        rgtPlate[1].tData.rgtCap[0].tFlag.tSelvedgeMachine.dDoneTrim1OpSide := 3, rgtPlate[1].tData.rgtCap[0].tFlag.tSelvedgeMachine.dDoneTrim2OppOpSide := 1, rgtPlate[1].tData.rgtCap[0].tFlag.tSelvedgeMachine.dDoneTrim3OppOpSide := 3, rgtPlate[2].tTracking.dPosition_cmm := 2104636, rgtPlate[2].tTracking.dPositionHead_cmm := 2234636, rgtPlate[2].tTracking.dPositionTail_cmm := 1974636, rgtPlate[2].tTracking.dLength_cmm := 260000, rgtPlate[2].tTracking.dIndexConvHead := 7, rgtPlate[2].tTracking.dIndexCapInConvHead := 2, rgtPlate[2].tTracking.dIndexConvTail := 6, rgtPlate[2].tTracking.dIndexCapInConvTail := 2, rgtPlate[2].tTracking.dLastConv := 6, rgtPlate[2].tTracking.dLastConvTail := 6, rgtPlate[2].tData.dLength_cmm := 260000, rgtPlate[2].tData.dTotalCaps := 1, rgtPlate[2].tData.rgtCap[0].dID := 4255236, rgtPlate[2].tData.rgtCap[0].dLength_cmm := 260000, rgtPlate[2].tData.rgtCap[0].dWidth_cmm := 360000, rgtPlate[2].tData.rgtCap[0].dThickness_cmm := 600, rgtPlate[2].tData.rgtCap[0].dFormat := 3, rgtPlate[2].tData.rgtCap[0].dNumLites := 2, rgtPlate[2].tData.rgtCap[0].dConvTotLength_cmm := 260000, rgtPlate[2].tData.rgtCap[0].dMinWidth_cmm := 360000, rgtPlate[2].tData.rgtCap[0].dMaxWidth_cmm := 360000, rgtPlate[2].tData.rgtCap[0].dGrossWidth_cmm := 377300, rgtPlate[2].tData.rgtCap[0].dDEdgeOpSide_cmm := 5000, rgtPlate[2].tData.rgtCap[0].dDEdgeOppOpSide_cmm := 5000, rgtPlate[2].tData.rgtCap[0].dCutWander_cmm := -3930, rgtPlate[2].tData.rgtCap[0].dNetWander_cmm := -6230, rgtPlate[2].tData.rgtCap[0].rgtLite[0].dID := 4255237, rgtPlate[2].tData.rgtCap[0].rgtLite[0].dProductionID := 1029, rgtPlate[2].tData.rgtCap[0].rgtLite[0].dQualityID := 10, rgtPlate[2].tData.rgtCap[0].rgtLite[0].dWidth_cmm := 180000, rgtPlate[2].tData.rgtCap[0].rgtLite[0].dBarycenter_cmm := -93930, rgtPlate[2].tData.rgtCap[0].rgtLite[1].dID := 4255238, rgtPlate[2].tData.rgtCap[0].rgtLite[1].dProductionID := 1029, rgtPlate[2].tData.rgtCap[0].rgtLite[1].dQualityID := 10, rgtPlate[2].tData.rgtCap[0].rgtLite[1].dWidth_cmm := 180000, rgtPlate[2].tData.rgtCap[0].rgtLite[1].dBarycenter_cmm := 86070, rgtPlate[2].tData.rgtCap[0].tFlag.xByYCut2 := 1, rgtPlate[2].tData.rgtCap[0].tFlag.xTrim2OpSide := 1, rgtPlate[2].tData.rgtCap[0].tFlag.xTrim1OpSide := 1, rgtPlate[2].tData.rgtCap[0].tFlag.xTrim1OppOpSide := 1, rgtPlate[2].tData.rgtCap[0].tFlag.xTrim2OppOpSide := 1, rgtPlate[2].tData.rgtCap[0].tFlag.rgxIntCut := 1, rgtPlate[2].tData.rgtCap[0].tFlag.xOptSelvedgeSel := 1, rgtPlate[2].tData.rgtCap[0].tFlag.xOptSplitBarSel := 1, rgtPlate[2].tData.rgtCap[0].tFlag.xOptSepRollSel := 1, rgtPlate[2].tData.rgtCap[0].tFlag.rgxXCutDoneHead := 2, rgtPlate[2].tData.rgtCap[0].tFlag.rgxXCutDoneTail := 2, rgtPlate[2].tData.rgtCap[0].tFlag.rgxYCutHeadDone := 835, rgtPlate[2].tData.rgtCap[0].tFlag.tSelvedgeMachine.dReqTrim2OpSide := 1, rgtPlate[2].tData.rgtCap[0].tFlag.tSelvedgeMachine.dReqTrim1OpSide := 3, rgtPlate[2].tData.rgtCap[0].tFlag.tSelvedgeMachine.dReqTrim1OppOpSide := 3, rgtPlate[2].tData.rgtCap[0].tFlag.tSelvedgeMachine.dReqTrim2OppOpSide := 1, rgtPlate[2].tData.rgtCap[0].tFlag.tSelvedgeMachine.dDoneTrim3OpSide := 3, rgtPlate[2].tData.rgtCap[0].tFlag.tSelvedgeMachine.dDoneTrim2OpSide := 1, rgtPlate[2].tData.rgtCap[0].tFlag.tSelvedgeMachine.dDoneTrim1OpSide := 3, rgtPlate[2].tData.rgtCap[0].tFlag.tSelvedgeMachine.dDoneTrim2OppOpSide := 1, rgtPlate[2].tData.rgtCap[0].tFlag.tSelvedgeMachine.dDoneTrim3OppOpSide := 3,
        rgtPlate[4].tTracking.dPosition_cmm := 1194845, rgtPlate[4].tTracking.dPositionHead_cmm := 1324845, rgtPlate[4].tTracking.dPositionTail_cmm := 1064845, rgtPlate[4].tTracking.dLength_cmm := 260000, rgtPlate[4].tTracking.dIndexConvHead := 5, rgtPlate[4].tTracking.dIndexCapInConvHead := 4, rgtPlate[4].tTracking.dIndexConvTail := 5, rgtPlate[4].tTracking.dIndexCapInConvTail := 4, rgtPlate[4].tTracking.dLastConv := 5, rgtPlate[4].tTracking.dLastConvTail := 5, rgtPlate[4].tData.dLength_cmm := 260000, rgtPlate[4].tData.dTotalCaps := 1, rgtPlate[4].tData.rgtCap[0].dID := 4255239, rgtPlate[4].tData.rgtCap[0].dLength_cmm := 260000, rgtPlate[4].tData.rgtCap[0].dWidth_cmm := 360000, rgtPlate[4].tData.rgtCap[0].dThickness_cmm := 600, rgtPlate[4].tData.rgtCap[0].dFormat := 2, rgtPlate[4].tData.rgtCap[0].dNumLites := 1, rgtPlate[4].tData.rgtCap[0].dConvTotLength_cmm := 260000, rgtPlate[4].tData.rgtCap[0].dMinWidth_cmm := 360000, rgtPlate[4].tData.rgtCap[0].dMaxWidth_cmm := 360000, rgtPlate[4].tData.rgtCap[0].dGrossWidth_cmm := 377400, rgtPlate[4].tData.rgtCap[0].dDEdgeOpSide_cmm := 5000, rgtPlate[4].tData.rgtCap[0].dDEdgeOppOpSide_cmm := 5000, rgtPlate[4].tData.rgtCap[0].dCutWander_cmm := -3930, rgtPlate[4].tData.rgtCap[0].dNetWander_cmm := -6130, rgtPlate[4].tData.rgtCap[0].rgtLite[0].dID := 4255240, rgtPlate[4].tData.rgtCap[0].rgtLite[0].dProductionID := 953, rgtPlate[4].tData.rgtCap[0].rgtLite[0].dQualityID := 10, rgtPlate[4].tData.rgtCap[0].rgtLite[0].dWidth_cmm := 360000, rgtPlate[4].tData.rgtCap[0].rgtLite[0].dBarycenter_cmm := -3930, rgtPlate[4].tData.rgtCap[0].tFlag.xByYCut2 := 1, rgtPlate[4].tData.rgtCap[0].tFlag.xTrim2OpSide := 1, rgtPlate[4].tData.rgtCap[0].tFlag.xTrim1OpSide := 1, rgtPlate[4].tData.rgtCap[0].tFlag.xTrim1OppOpSide := 1, rgtPlate[4].tData.rgtCap[0].tFlag.xTrim2OppOpSide := 1, rgtPlate[4].tData.rgtCap[0].tFlag.xOptSelvedgeSel := 1, rgtPlate[4].tData.rgtCap[0].tFlag.xOptSplitBarSel := 1, rgtPlate[4].tData.rgtCap[0].tFlag.xOptSepRollSel := 1, rgtPlate[4].tData.rgtCap[0].tFlag.rgxXCutDoneHead := 2, rgtPlate[4].tData.rgtCap[0].tFlag.rgxXCutDoneTail := 2, rgtPlate[4].tData.rgtCap[0].tFlag.rgxYCutHeadDone := 771, rgtPlate[4].tData.rgtCap[0].tFlag.tSelvedgeMachine.dReqTrim2OpSide := 1, rgtPlate[4].tData.rgtCap[0].tFlag.tSelvedgeMachine.dReqTrim1OpSide := 3, rgtPlate[4].tData.rgtCap[0].tFlag.tSelvedgeMachine.dReqTrim1OppOpSide := 3, rgtPlate[4].tData.rgtCap[0].tFlag.tSelvedgeMachine.dReqTrim2OppOpSide := 1, rgtPlate[4].tData.rgtCap[0].tFlag.tSelvedgeMachine.dDoneTrim2OpSide := 1, rgtPlate[4].tData.rgtCap[0].tFlag.tSelvedgeMachine.dDoneTrim2OppOpSide := 1, rgtPlate[5].tTracking.dPosition_cmm := 690000, rgtPlate[6].tTracking.dPosition_cmm := 306847, rgtPlate[6].tTracking.dPositionHead_cmm := 436847, rgtPlate[6].tTracking.dPositionTail_cmm := 176847, rgtPlate[6].tTracking.dLength_cmm := 260000, rgtPlate[6].tTracking.dIndexConvHead := 3, rgtPlate[6].tTracking.dIndexCapInConvHead := 6, rgtPlate[6].tTracking.dIndexConvTail := 2, rgtPlate[6].tTracking.dIndexCapInConvTail := 6, rgtPlate[6].tTracking.dLastConv := 3, rgtPlate[6].tTracking.dLastConvTail := 2, rgtPlate[6].tData.dLength_cmm := 260000,
        rgtPlate[6].tData.dTotalCaps := 1, rgtPlate[6].tData.rgtCap[0].dID := 4255241, rgtPlate[6].tData.rgtCap[0].dLength_cmm := 260000, rgtPlate[6].tData.rgtCap[0].dWidth_cmm := 360000, rgtPlate[6].tData.rgtCap[0].dThickness_cmm := 600, rgtPlate[6].tData.rgtCap[0].dFormat := 2, rgtPlate[6].tData.rgtCap[0].dNumLites := 1, rgtPlate[6].tData.rgtCap[0].dConvTotLength_cmm := 260000, rgtPlate[6].tData.rgtCap[0].dMinWidth_cmm := 360000, rgtPlate[6].tData.rgtCap[0].dMaxWidth_cmm := 360000, rgtPlate[6].tData.rgtCap[0].dGrossWidth_cmm := 377400, rgtPlate[6].tData.rgtCap[0].dDEdgeOpSide_cmm := 5000, rgtPlate[6].tData.rgtCap[0].dDEdgeOppOpSide_cmm := 5000, rgtPlate[6].tData.rgtCap[0].dCutWander_cmm := -3930, rgtPlate[6].tData.rgtCap[0].dNetWander_cmm := -6230, rgtPlate[6].tData.rgtCap[0].rgtLite[0].dID := 4255242, rgtPlate[6].tData.rgtCap[0].rgtLite[0].dProductionID := 953, rgtPlate[6].tData.rgtCap[0].rgtLite[0].dQualityID := 10, rgtPlate[6].tData.rgtCap[0].rgtLite[0].dWidth_cmm := 360000, rgtPlate[6].tData.rgtCap[0].rgtLite[0].dBarycenter_cmm := -3930, rgtPlate[6].tData.rgtCap[0].tFlag.xByYCut2 := 1, rgtPlate[6].tData.rgtCap[0].tFlag.xTrim2OpSide := 1, rgtPlate[6].tData.rgtCap[0].tFlag.xTrim1OpSide := 1, rgtPlate[6].tData.rgtCap[0].tFlag.xTrim1OppOpSide := 1, rgtPlate[6].tData.rgtCap[0].tFlag.xTrim2OppOpSide := 1, rgtPlate[6].tData.rgtCap[0].tFlag.xOptSelvedgeSel := 1, rgtPlate[6].tData.rgtCap[0].tFlag.xOptSplitBarSel := 1, rgtPlate[6].tData.rgtCap[0].tFlag.xOptSepRollSel := 1, rgtPlate[6].tData.rgtCap[0].tFlag.rgxXCutDoneHead := 2, rgtPlate[6].tData.rgtCap[0].tFlag.rgxXCutDoneTail := 2, rgtPlate[6].tData.rgtCap[0].tFlag.rgxYCutHeadDone := 771, rgtPlate[6].tData.rgtCap[0].tFlag.tSelvedgeMachine.dReqTrim2OpSide := 1, rgtPlate[6].tData.rgtCap[0].tFlag.tSelvedgeMachine.dReqTrim1OpSide := 3, rgtPlate[6].tData.rgtCap[0].tFlag.tSelvedgeMachine.dReqTrim1OppOpSide := 3, rgtPlate[6].tData.rgtCap[0].tFlag.tSelvedgeMachine.dReqTrim2OppOpSide := 1, rgtPlate[7].tTracking.dPosition_cmm := 3322205, rgtPlate[7].tTracking.dPositionHead_cmm := 3452205, rgtPlate[7].tTracking.dPositionTail_cmm := 3192205, rgtPlate[7].tTracking.dLength_cmm := 260000, rgtPlate[7].tTracking.dIndexConvHead := 11, rgtPlate[7].tTracking.dIndexCapInConvHead := 7, rgtPlate[7].tTracking.dIndexConvTail := 10, rgtPlate[7].tTracking.dIndexCapInConvTail := 7, rgtPlate[7].tTracking.dLastConv := 10, rgtPlate[7].tTracking.dLastConvTail := 10, rgtPlate[7].tData.dLength_cmm := 260000, rgtPlate[7].tData.dTotalCaps := 1, rgtPlate[7].tData.rgtCap[0].dID := 4255234, rgtPlate[7].tData.rgtCap[0].dLength_cmm := 260000, rgtPlate[7].tData.rgtCap[0].dWidth_cmm := 360000, rgtPlate[7].tData.rgtCap[0].dThickness_cmm := 600, rgtPlate[7].tData.rgtCap[0].dFormat := 2, rgtPlate[7].tData.rgtCap[0].dNumLites := 1, rgtPlate[7].tData.rgtCap[0].dConvTotLength_cmm := 260000, rgtPlate[7].tData.rgtCap[0].dMinWidth_cmm := 360000, rgtPlate[7].tData.rgtCap[0].dMaxWidth_cmm := 360000, rgtPlate[7].tData.rgtCap[0].dGrossWidth_cmm := 377400, rgtPlate[7].tData.rgtCap[0].dDEdgeOpSide_cmm := 5000, rgtPlate[7].tData.rgtCap[0].dDEdgeOppOpSide_cmm := 5000, rgtPlate[7].tData.rgtCap[0].dCutWander_cmm := -3930,
        rgtPlate[7].tData.rgtCap[0].dNetWander_cmm := -6130, rgtPlate[7].tData.rgtCap[0].rgtLite[0].dID := 4255235, rgtPlate[7].tData.rgtCap[0].rgtLite[0].dProductionID := 953, rgtPlate[7].tData.rgtCap[0].rgtLite[0].dQualityID := 10, rgtPlate[7].tData.rgtCap[0].rgtLite[0].dWidth_cmm := 360000, rgtPlate[7].tData.rgtCap[0].rgtLite[0].dBarycenter_cmm := -3930, rgtPlate[7].tData.rgtCap[0].tFlag.xByYCut2 := 1, rgtPlate[7].tData.rgtCap[0].tFlag.xTrim2OpSide := 1, rgtPlate[7].tData.rgtCap[0].tFlag.xTrim1OpSide := 1, rgtPlate[7].tData.rgtCap[0].tFlag.xTrim1OppOpSide := 1, rgtPlate[7].tData.rgtCap[0].tFlag.xTrim2OppOpSide := 1, rgtPlate[7].tData.rgtCap[0].tFlag.xOptSelvedgeSel := 1, rgtPlate[7].tData.rgtCap[0].tFlag.xOptSplitBarSel := 1, rgtPlate[7].tData.rgtCap[0].tFlag.xOptSepRollSel := 1, rgtPlate[7].tData.rgtCap[0].tFlag.xHookedGeom := 1, rgtPlate[7].tData.rgtCap[0].tFlag.rgxXCutDoneHead := 2, rgtPlate[7].tData.rgtCap[0].tFlag.rgxXCutDoneTail := 2, rgtPlate[7].tData.rgtCap[0].tFlag.rgxYCutHeadDone := 771, rgtPlate[7].tData.rgtCap[0].tFlag.tSelvedgeMachine.dReqTrim2OpSide := 1, rgtPlate[7].tData.rgtCap[0].tFlag.tSelvedgeMachine.dReqTrim1OpSide := 3, rgtPlate[7].tData.rgtCap[0].tFlag.tSelvedgeMachine.dReqTrim1OppOpSide := 3, rgtPlate[7].tData.rgtCap[0].tFlag.tSelvedgeMachine.dReqTrim2OppOpSide := 1, rgtPlate[7].tData.rgtCap[0].tFlag.tSelvedgeMachine.dDoneTrim3OpSide := 3, rgtPlate[7].tData.rgtCap[0].tFlag.tSelvedgeMachine.dDoneTrim2OpSide := 1, rgtPlate[7].tData.rgtCap[0].tFlag.tSelvedgeMachine.dDoneTrim1OpSide := 3, rgtPlate[7].tData.rgtCap[0].tFlag.tSelvedgeMachine.dDoneTrim2OppOpSide := 1, rgtPlate[7].tData.rgtCap[0].tFlag.tSelvedgeMachine.dDoneTrim3OppOpSide := 3); {access None}
   Z300_Conveyor : UDT_StandConv[29]; {access None}
        [0]   // M302M1
        [10]   // M305M1
        [21]   // M350M1
        [22]   // M310M1
        [1]   // M302M2
        [2]   // M302M3
        [3]   // M302M4
        [4]   // M302M5
        [8]   // M303M2
        [9]   // M304M1
        [5]   // M302M6
        [11]   // M306M1
        [7]   // M303M1
        [6]   // M302M7
        [12]   // M307AM1
        [13]   // M307AM2
        [14]   // M307AM3
        [15]   // M307AM4
        [16]   // M307BM1
        [17]   // M307CM1
        [18]   // M307DM1
        [19]   // M307EM1
        [20]   // M307FM1
        [23]   // M310M2
        [24]   // M310M3
        [25]   // M360M1
        [26]   // M315M1
        [27]   // M315M2
        [28]   // M315M3
   Z300_Conveyor_ALM : MAC_Conveyor_ZC_ALM[29]; {access Read Only}
        [5]   // M302M6
        [6]   // M302M7
        [0]   // M302M1
        [0].rgxStoppingFault_M[0].x2   // M302M1.Drive feedback error
        [0].rgxStoppingFault_M[0].x4   // M302M1.Motor thermal probe
        [0].rgxStoppingFault_M[0].x1   // M302M1.Drive error
        [0].rgxStoppingFault_M[0].x6   // M302M1.Drive not enabled
        [0].rgxStoppingFault_M[0].x0   // M302M1.Motor protection
        [0].rgxStoppingFault_M[0].x3   // M302M1.Local safety switch
        [0].rgxStoppingFault_M[0].x5   // M302M1.Braking resistor fault
        [14].rgxStoppingFault_M[0].x0   // M307AM3.Motor protection
        [10]   // M305M1
        [10].rgxStoppingFault_M[0].x2   // M305M1.Drive feedback error
        [10].rgxStoppingFault_M[0].x4   // M305M1.Motor thermal probe
        [10].rgxStoppingFault_M[0].x1   // M305M1.E76AZ1.Drive error
        [10].rgxStoppingFault_M[0].x6   // M305M1.Drive not enabled
        [10].rgxStoppingFault_M[0].x0   // M305M1.Motor protection
        [10].rgxStoppingFault_M[0].x3   // M305M1.Local safety switch
        [10].rgxStoppingFault_M[0].x5   // M305M1.Braking resistor fault
        [10].rgxFault_M[0].x0   // M313M3.E77QM1.Protection cooling fan
        [11].rgxStoppingFault_M[0].x2   // M306M1.Drive feedback error
        [11].rgxStoppingFault_M[0].x4   // M306M1.Motor thermal probe
        [11].rgxStoppingFault_M[0].x1   // M306M1.Drive error
        [11].rgxStoppingFault_M[0].x6   // M306M1.Drive not enabled
        [11].rgxStoppingFault_M[0].x0   // M306M1.Motor protection
        [11].rgxStoppingFault_M[0].x3   // M306M1.Local safety switch
        [11].rgxStoppingFault_M[0].x5   // M306M1.Braking resistor fault
        [17].rgxStoppingFault_M[0].x5   // M307CM1.Braking resistor fault
        [18].rgxStoppingFault_M[0].x2   // M307DM1.Drive feedback error
        [20].rgxStoppingFault_M[0].x0   // M307FM1.Protection motor
        [16].rgxStoppingFault_M[0].x0   // M307BM1.Protection motor
        [18].rgxStoppingFault_M[0].x1   // M307DM1.Drive error
        [21].rgxStoppingFault_M[0].x3   // M350M1.Local safety switch
        [16].rgxStoppingFault_M[0].x2   // M307BM1.Drive feedback error
        [12].rgxStoppingFault_M[0].x2   // M307AM1.Drive feedback error
        [12].rgxStoppingFault_M[0].x4   // M307AM1.Motor thermal probe
        [12].rgxStoppingFault_M[0].x1   // M307AM1.Drive error
        [12].rgxStoppingFault_M[0].x6   // M307AM1.Drive not enabled
        [21].rgxStoppingFault_M[0].x4   // M350M1.Motor thermal probe
        [16].rgxStoppingFault_M[0].x4   // M307BM1.Motor thermal probe
        [21]   // M350M1
        [13].rgxStoppingFault_M[0].x2   // M307AM2.Drive feedback error
        [13].rgxStoppingFault_M[0].x4   // M307AM2.Motor thermal probe
        [13].rgxStoppingFault_M[0].x1   // M307AM2.Drive error
        [13].rgxStoppingFault_M[0].x6   // M307AM2.Drive not enabled
        [15].rgxStoppingFault_M[0].x0   // M307AM4.Motor protection
        [15].rgxStoppingFault_M[0].x1   // M307AM4.Drive error
        [19].rgxStoppingFault_M[0].x2   // M307EM1.Drive feedback error
        [20].rgxStoppingFault_M[0].x2   // M307FM1.Drive feedback error
        [21].rgxStoppingFault_M[0].x1   // M350M1.Drive error
        [17].rgxStoppingFault_M[0].x0   // M307CM1.Protection motor
        [19].rgxStoppingFault_M[0].x1   // M307EM1.Drive error
        [22].rgxStoppingFault_M[0].x1   // M310M1.Drive error
        [17].rgxStoppingFault_M[0].x2   // M307CM1.Drive feedback error
        [22]   // M310M1
        [14].rgxStoppingFault_M[0].x2   // M307AM3.Drive feedback error
        [14].rgxStoppingFault_M[0].x4   // M307AM3.Motor thermal probe
        [14].rgxStoppingFault_M[0].x1   // M307AM3.Drive error
        [14].rgxStoppingFault_M[0].x6   // M307AM3.Drive not enabled
        [13].rgxStoppingFault_M[0].x0   // M307AM2.Motor protection
        [13].rgxStoppingFault_M[0].x3   // M307AM2.Local safety switch
        [18].rgxStoppingFault_M[0].x3   // M307DM1.Local safety switch
        [19].rgxStoppingFault_M[0].x3   // M307EM1.Local safety switch
        [22].rgxStoppingFault_M[0].x0   // M310M1.Protection motor
        [18].rgxStoppingFault_M[0].x0   // M307DM1.Protection motor
        [20].rgxStoppingFault_M[0].x1   // M307FM1.Drive error
        [22].rgxStoppingFault_M[0].x3   // M310M1.Local safety switch
        [17].rgxStoppingFault_M[0].x3   // M307CM1.Local safety switch
        [1]   // M302M2
        [1].rgxStoppingFault_M[0].x2   // M302M2.Drive feedback error
        [1].rgxStoppingFault_M[0].x4   // M302M2.Motor thermal probe
        [1].rgxStoppingFault_M[0].x1   // M302M2.Drive error
        [1].rgxStoppingFault_M[0].x6   // M302M2.Drive not enabled
        [1].rgxStoppingFault_M[0].x0   // M302M2.Motor protection
        [1].rgxStoppingFault_M[0].x3   // M302M2.Local safety switch
        [1].rgxStoppingFault_M[0].x5   // M302M2.Braking resistor fault
        [2]   // M302M3
        [2].rgxStoppingFault_M[0].x2   // M302M3.Drive feedback error
        [2].rgxStoppingFault_M[0].x4   // M302M3.Motor thermal probe
        [2].rgxStoppingFault_M[0].x1   // M302M3.Drive error
        [2].rgxStoppingFault_M[0].x6   // M302M3.Drive not enabled
        [2].rgxStoppingFault_M[0].x0   // M302M3.Motor protection
        [2].rgxStoppingFault_M[0].x3   // M302M3.Local safety switch
        [2].rgxStoppingFault_M[0].x5   // M302M3.Braking resistor fault
        [3]   // M302M4
        [3].rgxStoppingFault_M[0].x2   // M302M4.Drive feedback error
        [3].rgxStoppingFault_M[0].x4   // M302M4.Motor thermal probe
        [3].rgxStoppingFault_M[0].x1   // M302M4.Drive error
        [3].rgxStoppingFault_M[0].x6   // M302M4.Drive not enabled
        [3].rgxStoppingFault_M[0].x0   // M302M4.Motor protection
        [3].rgxStoppingFault_M[0].x3   // M302M4.Local safety switch
        [3].rgxStoppingFault_M[0].x5   // M302M4.Braking resistor fault
        [4]   // M302M5
        [4].rgxStoppingFault_M[0].x2   // M302M5.Drive feedback error
        [4].rgxStoppingFault_M[0].x4   // M302M5.Motor thermal probe
        [4].rgxStoppingFault_M[0].x1   // M302M5.Drive error
        [4].rgxStoppingFault_M[0].x6   // M302M5.Drive not enabled
        [4].rgxStoppingFault_M[0].x0   // M302M5.Motor protection
        [4].rgxStoppingFault_M[0].x3   // M302M5.Local safety switch
        [4].rgxStoppingFault_M[0].x5   // M302M5.Braking resistor fault
        [5].rgxStoppingFault_M[0].x2   // M302M6.Drive feedback error
        [5].rgxStoppingFault_M[0].x4   // M302M6.Motor thermal probe
        [5].rgxStoppingFault_M[0].x1   // M302M6.Drive error
        [5].rgxStoppingFault_M[0].x6   // M302M6.Drive not enabled
        [5].rgxStoppingFault_M[0].x0   // M302M6.Motor protection
        [5].rgxStoppingFault_M[0].x3   // M302M6.Local safety switch
        [5].rgxStoppingFault_M[0].x5   // M302M6.Braking resistor fault
        [16].rgxStoppingFault_M[0].x5   // M307BM1.Braking resistor fault
        [17].rgxStoppingFault_M[0].x4   // M307CM1.Motor thermal probe
        [21].rgxStoppingFault_M[0].x0   // M350M1.Protection motor
        [17].rgxStoppingFault_M[0].x1   // M307CM1.Drive error
        [16].rgxStoppingFault_M[0].x1   // M307BM1.Drive error
        [19].rgxStoppingFault_M[0].x0   // M307EM1.Protection motor
        [16].rgxStoppingFault_M[0].x3   // M307BM1.Local safety switch
        [6].rgxStoppingFault_M[0].x2   // M302M7.Drive feedback error
        [6].rgxStoppingFault_M[0].x4   // M302M7.Motor thermal probe
        [6].rgxStoppingFault_M[0].x1   // M302M7.Drive error
        [6].rgxStoppingFault_M[0].x6   // M302M7.Drive not enabled
        [6].rgxStoppingFault_M[0].x0   // M302M7.Motor protection
        [6].rgxStoppingFault_M[0].x3   // M302M7.Local safety switch
        [6].rgxStoppingFault_M[0].x5   // M302M7.Braking resistor fault
        [6].rgxFault_M[0].x0   // M311M1.E70QM1.Protection cooling fan
        [7].rgxStoppingFault_M[0].x2   // M303M1.Drive feedback error
        [7].rgxStoppingFault_M[0].x4   // M303M1.Motor thermal probe
        [7].rgxStoppingFault_M[0].x1   // M303M1.Drive error
        [7].rgxStoppingFault_M[0].x6   // M303M1.Drive not enabled
        [7].rgxStoppingFault_M[0].x0   // M303M1.Motor protection
        [7].rgxStoppingFault_M[0].x3   // M303M1.Local safety switch
        [7].rgxStoppingFault_M[0].x5   // M303M1.Braking resistor fault
        [7].rgxFault_M[0].x0   // M312M1.E73QM1.Protection cooling fan
        [8]   // M303M2
        [8].rgxStoppingFault_M[0].x2   // M303M2.Drive feedback error
        [8].rgxStoppingFault_M[0].x4   // M303M2.Motor thermal probe
        [8].rgxStoppingFault_M[0].x1   // M303M2.Drive error
        [8].rgxStoppingFault_M[0].x6   // M303M2.Drive not enabled
        [8].rgxStoppingFault_M[0].x0   // M303M2.Motor protection
        [8].rgxStoppingFault_M[0].x3   // M303M2.Local safety switch
        [8].rgxStoppingFault_M[0].x5   // M303M2.Braking resistor fault
        [8].rgxFault_M[0].x0   // M313M1.E74QM1.Protection cooling fan
        [9]   // M304M1
        [9].rgxStoppingFault_M[0].x2   // M304M1.Drive feedback error
        [9].rgxStoppingFault_M[0].x4   // M304M1.Motor thermal probe
        [9].rgxStoppingFault_M[0].x1   // M304M1.Drive error
        [9].rgxStoppingFault_M[0].x6   // M304M1.Drive not enabled
        [9].rgxStoppingFault_M[0].x0   // M304M1.Motor protection
        [9].rgxStoppingFault_M[0].x3   // M304M1.Local safety switch
        [9].rgxStoppingFault_M[0].x5   // M304M1.Braking resistor fault
        [9].rgxFault_M[0].x0   // M313M2.E76QM1.Protection cooling fan
        [7]   // M303M1
        [11]   // M306M1
        [12]   // M307AM1
        [13]   // M307AM2
        [14]   // M307AM3
        [15]   // M307AM4
        [16]   // M307BM1
        [17]   // M307CM1
        [18]   // M307DM1
        [19]   // M307EM1
        [20]   // M307FM1
        [23]   // M310M2
        [24]   // M310M3
        [25]   // M360M1
        [26]   // M315M1
        [27]   // M315M2
        [28]   // M315M3
        [14].rgxStoppingFault_M[0].x3   // M307AM3.Local safety switch
        [14].rgxStoppingFault_M[0].x5   // M307AM3.Braking resistor fault
        [13].rgxStoppingFault_M[0].x5   // M307AM2.Braking resistor fault
        [15].rgxStoppingFault_M[0].x2   // M307AM4.Drive feedback error
        [15].rgxStoppingFault_M[0].x3   // M307AM4.Local safety switch
        [15].rgxStoppingFault_M[0].x4   // M307AM4.Motor thermal probe
        [15].rgxStoppingFault_M[0].x5   // M307AM4.Braking resistor fault
        [12].rgxStoppingFault_M[0].x0   // M307AM1.Motor protection
        [12].rgxStoppingFault_M[0].x3   // M307AM1.Local safety switch
        [12].rgxStoppingFault_M[0].x5   // M307AM1.Braking resistor fault
        [20].rgxStoppingFault_M[0].x3   // M307FM1.Local safety switch
        [18].rgxStoppingFault_M[0].x4   // M307DM1.Motor thermal probe
        [19].rgxStoppingFault_M[0].x4   // M307EM1.Motor thermal probe
        [20].rgxStoppingFault_M[0].x4   // M307FM1.Motor thermal probe
        [18].rgxStoppingFault_M[0].x5   // M307DM1.Braking resistor fault
        [19].rgxStoppingFault_M[0].x5   // M307EM1.Braking resistor fault
        [20].rgxStoppingFault_M[0].x5   // M307FM1.Braking resistor fault
        [21].rgxStoppingFault_M[0].x2   // M350M1.Drive feedback error
        [22].rgxStoppingFault_M[0].x2   // M310M1.Drive feedback error
        [21].rgxStoppingFault_M[0].x5   // M350M1 Braking resistor fault
        [22].rgxStoppingFault_M[0].x4   // M310M1.Motor thermal probe
        [22].rgxStoppingFault_M[0].x5   // M310M1.Braking resistor fault
        [23].rgxStoppingFault_M[0].x0   // M310M2.Protection motor
        [23].rgxStoppingFault_M[0].x1   // M310M2.Drive error
        [23].rgxStoppingFault_M[0].x2   // M310M2.Drive feedback error
        [23].rgxStoppingFault_M[0].x3   // M310M2.Local safety switch
        [23].rgxStoppingFault_M[0].x4   // M310M2.Motor thermal probe
        [23].rgxStoppingFault_M[0].x5   // M310M2.Braking resistor fault
        [24].rgxStoppingFault_M[0].x0   // M310M3.Protection motor
        [24].rgxStoppingFault_M[0].x1   // M310M3.Drive error
        [24].rgxStoppingFault_M[0].x2   // M310M3.Drive feedback error
        [24].rgxStoppingFault_M[0].x3   // M310M3.Local safety switch
        [24].rgxStoppingFault_M[0].x4   // M310M3.Motor thermal probe
        [24].rgxStoppingFault_M[0].x5   // M310M3.Braking resistor fault
        [25].rgxStoppingFault_M[0].x0   // M360M1.Protection motor
        [25].rgxStoppingFault_M[0].x1   // M360M1.Drive error
        [25].rgxStoppingFault_M[0].x2   // M360M1.Drive feedback error
        [25].rgxStoppingFault_M[0].x3   // M360M1.Local safety switch
        [25].rgxStoppingFault_M[0].x4   // M360M1.Motor thermal probe
        [25].rgxStoppingFault_M[0].x5   // M360M1.Braking resistor fault
        [26].rgxStoppingFault_M[0].x0   // M315M1.Protection motor
        [26].rgxStoppingFault_M[0].x1   // M315M1.Drive error
        [26].rgxStoppingFault_M[0].x2   // M315M1.Drive feedback error
        [26].rgxStoppingFault_M[0].x3   // M315M1.Local safety switch
        [26].rgxStoppingFault_M[0].x4   // M315M1.Motor thermal probe
        [26].rgxStoppingFault_M[0].x5   // M315M1.Braking resistor fault
        [27].rgxStoppingFault_M[0].x0   // M315M2.Protection motor
        [28].rgxStoppingFault_M[0].x0   // M315M3.Protection motor
        [27].rgxStoppingFault_M[0].x1   // M315M2.Drive error
        [28].rgxStoppingFault_M[0].x1   // M315M3.Drive error
        [27].rgxStoppingFault_M[0].x2   // M315M2.Drive feedback error
        [28].rgxStoppingFault_M[0].x2   // M315M3.Drive feedback error
        [27].rgxStoppingFault_M[0].x3   // M315M2.Local safety switch
        [28].rgxStoppingFault_M[0].x3   // M315M3.Local safety switch
        [27].rgxStoppingFault_M[0].x4   // M315M2.Motor thermal probe
        [28].rgxStoppingFault_M[0].x4   // M315M3.Motor thermal probe
        [27].rgxStoppingFault_M[0].x5   // M315M2.Braking resistor fault
        [28].rgxStoppingFault_M[0].x5   // M315M3.Braking resistor fault
   Z300_Conveyor_Conf : UDT_Conveyor_Config[29] := ([0].dLengthConveyor_cmm := 37500, [0].dWidthConveyor_cmm := 450000, [0].dPitchRoller := 25000, [0].dZoneConveyor := 1, [0].dIndexMainSpeed := 1, [0].xContinuousConveyor := 1, [0].rAccH_ms2 := 1.2, [0].rDecH_ms2 := 1.2, [0].rAccH_s := 0.75, [0].rDecH_s := 0.75, [0].rAccL_ms2 := 0.7, [0].rDecL_ms2 := 0.7, [0].rAccL_s := 1.29, [0].rDecL_s := 1.29, [0].rgxAllowedCullet := 16777216, [0].rgxAllowedQuality := 536870912, [1].dLengthConveyor_cmm := 50000, [1].dWidthConveyor_cmm := 450000, [1].dPitchRoller := 25000, [1].dMachineIndex := 1, [1].dZoneConveyor := 1, [1].dIndexMainSpeed := 1, [1].xContinuousConveyor := 1, [1].rAccH_ms2 := 1.2, [1].rDecH_ms2 := 1.2, [1].rAccH_s := 0.75, [1].rDecH_s := 0.75, [1].rAccL_ms2 := 0.7, [1].rDecL_ms2 := 0.7, [1].rAccL_s := 1.29, [1].rDecL_s := 1.29, [1].rgxAllowedCullet := 16777216, [1].rgxAllowedQuality := 536870912, [2].dLengthConveyor_cmm := 125000, [2].dWidthConveyor_cmm := 450000, [2].dPitchRoller := 25000, [2].dMachineIndex := 2, [2].dZoneConveyor := 1, [2].dIndexMainSpeed := 1, [2].xContinuousConveyor := 1, [2].rAccH_ms2 := 1.2, [2].rDecH_ms2 := 1.2, [2].rAccH_s := 0.75, [2].rDecH_s := 0.75, [2].rAccL_ms2 := 0.7, [2].rDecL_ms2 := 0.7, [2].rAccL_s := 1.29, [2].rDecL_s := 1.29, [2].rgxAllowedCullet := 16777216, [2].rgxAllowedQuality := 536870912, [3].dLengthConveyor_cmm := 250000, [3].dWidthConveyor_cmm := 450000, [3].dPitchRoller := 25000, [3].dMachineIndex := 3, [3].dZoneConveyor := 1, [3].dIndexMainSpeed := 1, [3].xContinuousConveyor := 1, [3].rAccH_ms2 := 1.2, [3].rDecH_ms2 := 1.2, [3].rAccH_s := 0.75,
        [3].rDecH_s := 0.75, [3].rAccL_ms2 := 0.7, [3].rDecL_ms2 := 0.7, [3].rAccL_s := 1.29, [3].rDecL_s := 1.29, [3].rgxAllowedCullet := 16777216, [3].rgxAllowedQuality := 536870912, [4].dLengthConveyor_cmm := 250000, [4].dWidthConveyor_cmm := 450000, [4].dPitchRoller := 25000, [4].dMachineIndex := 4, [4].dZoneConveyor := 1, [4].dIndexMainSpeed := 1, [4].xContinuousConveyor := 1, [4].rAccH_ms2 := 1.2, [4].rDecH_ms2 := 1.2, [4].rAccH_s := 0.75, [4].rDecH_s := 0.75, [4].rAccL_ms2 := 0.7, [4].rDecL_ms2 := 0.7, [4].rAccL_s := 1.29, [4].rDecL_s := 1.29, [4].rgxAllowedCullet := 16777216, [4].rgxAllowedQuality := 536870912, [5].dLengthConveyor_cmm := 914500, [5].dWidthConveyor_cmm := 450000, [5].dPitchRoller := 25000, [5].dMachineIndex := 5, [5].dZoneConveyor := 1, [5].dMotorNumber := 1, [5].dIndexMainSpeed := 3, [5].xContinuousConveyor := 1, [5].rAccH_ms2 := 1.2, [5].rDecH_ms2 := 1.2, [5].rAccH_s := 0.75, [5].rDecH_s := 0.75, [5].rAccL_ms2 := 0.7, [5].rDecL_ms2 := 0.7, [5].rAccL_s := 1.29, [5].rDecL_s := 1.29, [5].rgxAllowedCullet := 16777216, [5].rgxAllowedQuality := 536870912, [6].dLengthConveyor_cmm := 500000, [6].dWidthConveyor_cmm := 450000, [6].dPitchRoller := 25000, [6].dMachineIndex := 6, [6].dZoneConveyor := 1, [6].dIndexMainSpeed := 3, [6].xContinuousConveyor := 1, [6].rAccH_ms2 := 1.2, [6].rDecH_ms2 := 1.2, [6].rAccH_s := 0.75, [6].rDecH_s := 0.75, [6].rAccL_ms2 := 0.7, [6].rDecL_ms2 := 0.7, [6].rAccL_s := 1.29, [6].rDecL_s := 1.29, [6].rgxAllowedCullet := 16777216, [6].rgxAllowedQuality := 536870912, [7].dLengthConveyor_cmm := 500000,
        [7].dWidthConveyor_cmm := 450000, [7].dPitchRoller := 25000, [7].dMachineIndex := 7, [7].dZoneConveyor := 1, [7].dIndexMainSpeed := 3, [7].xContinuousConveyor := 1, [7].rAccH_ms2 := 1.2, [7].rDecH_ms2 := 1.2, [7].rAccH_s := 0.75, [7].rDecH_s := 0.75, [7].rAccL_ms2 := 0.7, [7].rDecL_ms2 := 0.7, [7].rAccL_s := 1.29, [7].rDecL_s := 1.29, [7].rgxAllowedCullet := 16777216, [7].rgxAllowedQuality := 536870912, [8].dLengthConveyor_cmm := 75000, [8].dWidthConveyor_cmm := 450000, [8].dPitchRoller := 25000, [8].dMachineIndex := 8, [8].dZoneConveyor := 1, [8].dIndexMainSpeed := 3, [8].xContinuousConveyor := 1, [8].rAccH_ms2 := 1.2, [8].rDecH_ms2 := 1.2, [8].rAccH_s := 1.25, [8].rDecH_s := 1.25, [8].rAccL_ms2 := 0.7, [8].rDecL_ms2 := 0.7, [8].rAccL_s := 2.14, [8].rDecL_s := 2.14, [8].rgxAllowedCullet := 16777216, [8].rgxAllowedQuality := 536870912, [9].dLengthConveyor_cmm := 325000, [9].dWidthConveyor_cmm := 450000, [9].dPitchRoller := 25000, [9].dMachineIndex := 9, [9].dZoneConveyor := 1, [9].dIndexMainSpeed := 3, [9].xContinuousConveyor := 1, [9].rAccH_ms2 := 1.2, [9].rDecH_ms2 := 1.2, [9].rAccH_s := 1.25, [9].rDecH_s := 1.25, [9].rAccL_ms2 := 0.7, [9].rDecL_ms2 := 0.7, [9].rAccL_s := 2.14, [9].rDecL_s := 2.14, [9].rgxAllowedCullet := 16777216, [9].rgxAllowedQuality := 536870912, [10].dLengthConveyor_cmm := 400000, [10].dWidthConveyor_cmm := 450000, [10].dPitchRoller := 25000, [10].dMachineIndex := 10, [10].dZoneConveyor := 1, [10].dIndexMainSpeed := 3, [10].xContinuousConveyor := 1, [10].rAccH_ms2 := 1.2, [10].rDecH_ms2 := 1.2, [10].rAccH_s := 1.25,
        [10].rDecH_s := 1.25, [10].rAccL_ms2 := 0.7, [10].rDecL_ms2 := 0.7, [10].rAccL_s := 2.14, [10].rDecL_s := 2.14, [10].rgxAllowedCullet := 16777216, [10].rgxAllowedQuality := 536870912, [11].dLengthConveyor_cmm := 350000, [11].dWidthConveyor_cmm := 450000, [11].dPitchRoller := 25000, [11].dMachineIndex := 11, [11].dZoneConveyor := 1, [11].dMotorNumber := 1, [11].xContinuousConveyor := 1, [11].rAccH_ms2 := 1.2, [11].rDecH_ms2 := 1.2, [11].rAccH_s := 1.25, [11].rDecH_s := 1.25, [11].rAccL_ms2 := 0.7, [11].rDecL_ms2 := 0.7, [11].rAccL_s := 2.14, [11].rDecL_s := 2.14, [11].rgxAllowedCullet := 16777216, [11].rgxAllowedQuality := 536870912, [12].dLengthConveyor_cmm := 450000, [12].dWidthConveyor_cmm := 450000, [12].dPitchRoller := 25000, [12].dMachineIndex := 12, [12].dZoneConveyor := 2, [12].dSpaceRestartPlate_cmm := 150000, [12].xWaitGlassForStop := 1, [12].rAccH_ms2 := 1.2, [12].rDecH_ms2 := 1.2, [12].rAccH_s := 1.25, [12].rDecH_s := 1.25, [12].rAccL_ms2 := 0.7, [12].rDecL_ms2 := 0.7, [12].rAccL_s := 2.14, [12].rDecL_s := 2.14, [12].rgxAllowedCullet := 16777216, [12].rgxAllowedQuality := 536870912, [13].dLengthConveyor_cmm := 300000, [13].dWidthConveyor_cmm := 450000, [13].dPitchRoller := 25000, [13].dMachineIndex := 13, [13].dZoneConveyor := 2, [13].dMotorNumber := 1, [13].dSpaceRestartPlate_cmm := 150000, [13].xWaitGlassForStop := 1, [13].rAccH_ms2 := 1.2, [13].rDecH_ms2 := 1.2, [13].rAccH_s := 1.25, [13].rDecH_s := 1.25, [13].rAccL_ms2 := 0.7, [13].rDecL_ms2 := 0.7, [13].rAccL_s := 2.14, [13].rDecL_s := 2.14, [13].rgxAllowedCullet := 16777216, [13].rgxAllowedQuality := 536870912, [14].dLengthConveyor_cmm := 100000,
